   // TANK_CONTROL_1S.PVVX_OUT_DATA.PVVB_DemandsCompleted[10] := False;
   // TANK_CONTROL_1S.PVVX_OUT_DATA.PVVB_DemandsCompleted[9] := False;
   // TANK_CONTROL_1S.PVVX_OUT_DATA.PVVB_DemandsCompleted[8] := False;
   // TANK_CONTROL_1S.PVVX_OUT_DATA.PVVB_DemandsCompleted[7] := False;
   // TANK_CONTROL_1S.PVVX_OUT_DATA.PVVB_DemandsCompleted[6] := False;
   // TANK_CONTROL_1S.PVVX_OUT_DATA.PVVB_DemandsCompleted[5] := False;
   // TANK_CONTROL_6P.DWELL_TIMER.IN := False;
   // TANK_CONTROL_6P.MONITOR_TIMER.IN := False;
   // TANK_CONTROL_6P.ReOx_InitialTargetpHLevelAchieved := False;
   // TANK_CONTROL_1S.PVVX_OUT_DATA.PVVB_DemandsCompleted[4] := False;
   // TANK_CONTROL_1S.PVVX_OUT_DATA.PVVB_DemandsCompleted[3] := False;
   // TANK_CONTROL_1S.PVVX_OUT_DATA.PVVB_DemandsCompleted[2] := False;
   // TANK_CONTROL_1S.PVVX_OUT_DATA.PVVB_DemandsCompleted[1] := False;
   // TANK_CONTROL_1S.PVVX_OUT_DATA.PVVA_Alarms[14] := False;
   // TANK_CONTROL_1S.PVVX_OUT_DATA.PVVA_Alarms[13] := False;
   // TANK_CONTROL_1S.PVVX_OUT_DATA.PVVA_Alarms[12] := False;
   // TANK_CONTROL_1S.PVVX_OUT_DATA.PVVA_Alarms[11] := False;
   // TANK_CONTROL_1S.PVVX_OUT_DATA.PVVA_Alarms[10] := False;
   // TANK_CONTROL_1S.PVVX_OUT_DATA.PVVA_Alarms[9] := False;
   // TANK_CONTROL_1S.PVVX_OUT_DATA.PVVA_Alarms[8] := False;
   // TANK_CONTROL_1S.PVVX_OUT_DATA.PVVA_Alarms[7] := False;
   // TANK_CONTROL_1S.PVVX_OUT_DATA.PVVA_Alarms[6] := False;
   // TANK_CONTROL_1S.PVVX_OUT_DATA.PVVA_Alarms[5] := False;
   // TANK_CONTROL_1S.PVVX_OUT_DATA.PVVA_Alarms[4] := False;
   // TANK_CONTROL_1S.PVVX_OUT_DATA.PVVA_Alarms[3] := False;
   // TANK_CONTROL_1S.PVVX_OUT_DATA.PVVA_Alarms[2] := False;
   // TANK_CONTROL_1S.PVVX_OUT_DATA.PVVA_Alarms[1] := False;
   // TANK_CONTROL_1S.PVVX_OUT_DATA.PVVA_DemandsCompleted[14] := False;
   // TANK_CONTROL_1S.PVVX_OUT_DATA.PVVA_DemandsCompleted[13] := False;
   // TANK_CONTROL_1S.PVVX_OUT_DATA.PVVA_DemandsCompleted[12] := False;
   // TANK_CONTROL_1S.PVVX_OUT_DATA.PVVA_DemandsCompleted[11] := False;
   // TANK_CONTROL_1S.PVVX_OUT_DATA.PVVA_DemandsCompleted[10] := False;
   // TANK_CONTROL_1S.PVVX_OUT_DATA.PVVA_DemandsCompleted[9] := False;
   // TANK_CONTROL_1S.PVVX_OUT_DATA.PVVA_DemandsCompleted[8] := False;
   // TANK_CONTROL_1S.PVVX_OUT_DATA.PVVA_DemandsCompleted[7] := False;
   // TANK_CONTROL_1S.PVVX_OUT_DATA.PVVA_DemandsCompleted[6] := False;
   // TANK_CONTROL_1S.PVVX_OUT_DATA.PVVA_DemandsCompleted[5] := False;
   // TANK_CONTROL_1S.PVVX_OUT_DATA.PVVA_DemandsCompleted[4] := False;
   // TANK_CONTROL_1S.PVVX_OUT_DATA.PVVA_DemandsCompleted[3] := False;
   // TANK_CONTROL_1S.PVVX_OUT_DATA.PVVA_DemandsCompleted[2] := False;
   // TANK_CONTROL_1S.PVVX_OUT_DATA.PVVA_DemandsCompleted[1] := False;
   // TANK_CONTROL_1P.GTT_OUT_DATA.GTT_Alarms[14] := False;
   // TANK_CONTROL_1P.GTT_OUT_DATA.GTT_Alarms[13] := False;
   // TANK_CONTROL_1P.GTT_OUT_DATA.GTT_Alarms[12] := False;
   // TANK_CONTROL_1P.GTT_OUT_DATA.GTT_Alarms[11] := False;
   // TANK_CONTROL_1P.GTT_OUT_DATA.GTT_Alarms[10] := False;
   // TANK_CONTROL_1P.GTT_OUT_DATA.GTT_Alarms[9] := False;
   // TANK_CONTROL_1P.GTT_OUT_DATA.GTT_Alarms[8] := False;
   // TANK_CONTROL_1P.GTT_OUT_DATA.GTT_Alarms[7] := False;
   // TANK_CONTROL_1P.GTT_OUT_DATA.GTT_Alarms[6] := False;
   // TANK_CONTROL_1P.GTT_OUT_DATA.GTT_Alarms[5] := False;
   // TANK_CONTROL_1P.GTT_OUT_DATA.GTT_Alarms[4] := False;
   // TANK_CONTROL_1P.GTT_OUT_DATA.GTT_Alarms[3] := False;
   // TANK_CONTROL_1P.GTT_OUT_DATA.GTT_Alarms[2] := False;
   // TANK_CONTROL_1P.GTT_OUT_DATA.GTT_Alarms[1] := False;
   // TANK_CONTROL_1P.GTT_OUT_DATA.GTT_DemandsCompleted[14] := False;
   // TANK_CONTROL_1P.GTT_OUT_DATA.GTT_DemandsCompleted[13] := False;
   // TANK_CONTROL_1P.GTT_OUT_DATA.GTT_DemandsCompleted[12] := False;
   // TANK_CONTROL_1P.GTT_OUT_DATA.GTT_DemandsCompleted[11] := False;
   // TANK_CONTROL_1P.GTT_OUT_DATA.GTT_DemandsCompleted[10] := False;
   // TANK_CONTROL_1P.GTT_OUT_DATA.GTT_DemandsCompleted[9] := False;
   // TANK_CONTROL_1P.GTT_OUT_DATA.GTT_DemandsCompleted[8] := False;
   // TANK_CONTROL_1P.GTT_OUT_DATA.GTT_DemandsCompleted[7] := False;
   // TANK_CONTROL_1P.GTT_OUT_DATA.GTT_DemandsCompleted[6] := False;
   // TANK_CONTROL_1P.GTT_OUT_DATA.GTT_DemandsCompleted[5] := False;
   // TANK_CONTROL_1P.GTT_OUT_DATA.GTT_DemandsCompleted[4] := False;
   // TANK_CONTROL_1P.GTT_OUT_DATA.GTT_DemandsCompleted[3] := False;
   // TANK_CONTROL_1P.GTT_OUT_DATA.GTT_DemandsCompleted[2] := False;
   // TANK_CONTROL_1P.GTT_OUT_DATA.GTT_DemandsCompleted[1] := False;
   // TANK_CONTROL_1P.PVVX_OUT_DATA.PVVB_Alarms[14] := False;
   // TANK_CONTROL_1P.PVVX_OUT_DATA.PVVB_Alarms[13] := False;
   // TANK_CONTROL_1P.PVVX_OUT_DATA.PVVB_Alarms[12] := False;
   // TANK_CONTROL_1P.PVVX_OUT_DATA.PVVB_Alarms[11] := False;
   // TANK_CONTROL_1P.PVVX_OUT_DATA.PVVB_Alarms[10] := False;
   // TANK_CONTROL_1P.PVVX_OUT_DATA.PVVB_Alarms[9] := False;
   // TANK_CONTROL_1P.PVVX_OUT_DATA.PVVB_Alarms[8] := False;
   // TANK_CONTROL_1P.PVVX_OUT_DATA.PVVB_Alarms[7] := False;
   // TANK_CONTROL_1P.PVVX_OUT_DATA.PVVB_Alarms[6] := False;
   // TANK_CONTROL_1P.PVVX_OUT_DATA.PVVB_Alarms[5] := False;
   // TANK_CONTROL_1P.PVVX_OUT_DATA.PVVB_Alarms[4] := False;
   // TANK_CONTROL_1P.PVVX_OUT_DATA.PVVB_Alarms[3] := False;
   // TANK_CONTROL_1P.PVVX_OUT_DATA.PVVB_Alarms[2] := False;
   // TANK_CONTROL_1P.PVVX_OUT_DATA.PVVB_Alarms[1] := False;
   // TANK_CONTROL_1P.PVVX_OUT_DATA.PVVB_DemandsCompleted[14] := False;
   // TANK_CONTROL_1P.PVVX_OUT_DATA.PVVB_DemandsCompleted[13] := False;
   // TANK_CONTROL_1P.PVVX_OUT_DATA.PVVB_DemandsCompleted[12] := False;
   // TANK_CONTROL_1P.PVVX_OUT_DATA.PVVB_DemandsCompleted[11] := False;
   // TANK_CONTROL_1P.PVVX_OUT_DATA.PVVB_DemandsCompleted[10] := False;
   // TANK_CONTROL_1P.PVVX_OUT_DATA.PVVB_DemandsCompleted[9] := False;
   // TANK_CONTROL_1P.PVVX_OUT_DATA.PVVB_DemandsCompleted[8] := False;
   // TANK_CONTROL_1P.PVVX_OUT_DATA.PVVB_DemandsCompleted[7] := False;
   // TANK_CONTROL_1P.PVVX_OUT_DATA.PVVB_DemandsCompleted[6] := False;
   // TANK_CONTROL_1P.PVVX_OUT_DATA.PVVB_DemandsCompleted[5] := False;
   // TANK_CONTROL_1P.PVVX_OUT_DATA.PVVB_DemandsCompleted[4] := False;
   // TANK_CONTROL_1P.PVVX_OUT_DATA.PVVB_DemandsCompleted[3] := False;
   // TANK_CONTROL_1P.PVVX_OUT_DATA.PVVB_DemandsCompleted[2] := False;
   // TANK_CONTROL_1P.PVVX_OUT_DATA.PVVB_DemandsCompleted[1] := False;
   // TANK_CONTROL_1P.PVVX_OUT_DATA.PVVA_Alarms[14] := False;
   // TANK_CONTROL_1P.PVVX_OUT_DATA.PVVA_Alarms[13] := False;
   // TANK_CONTROL_1P.PVVX_OUT_DATA.PVVA_Alarms[12] := False;
   // TANK_CONTROL_1P.PVVX_OUT_DATA.PVVA_Alarms[11] := False;
   // TANK_CONTROL_1P.PVVX_OUT_DATA.PVVA_Alarms[10] := False;
   // TANK_CONTROL_1P.PVVX_OUT_DATA.PVVA_Alarms[9] := False;
   // TANK_CONTROL_1P.PVVX_OUT_DATA.PVVA_Alarms[8] := False;
   // TANK_CONTROL_1P.PVVX_OUT_DATA.PVVA_Alarms[7] := False;
   // TANK_CONTROL_1P.PVVX_OUT_DATA.PVVA_Alarms[6] := False;
   // TANK_CONTROL_1P.PVVX_OUT_DATA.PVVA_Alarms[5] := False;
   // TANK_CONTROL_1P.PVVX_OUT_DATA.PVVA_Alarms[4] := False;
   // TANK_CONTROL_1P.PVVX_OUT_DATA.PVVA_Alarms[3] := False;
   // TANK_CONTROL_6S.DWELL_TIMER.IN := False;
   // TANK_CONTROL_6S.MONITOR_TIMER.IN := False;
   // TANK_CONTROL_6S.ReOx_InitialTargetpHLevelAchieved := False;
   // TANK_CONTROL_1P.PVVX_OUT_DATA.PVVA_Alarms[2] := False;
   // TANK_CONTROL_1P.PVVX_OUT_DATA.PVVA_Alarms[1] := False;
   // TANK_CONTROL_1P.PVVX_OUT_DATA.PVVA_DemandsCompleted[14] := False;
   // TANK_CONTROL_1P.PVVX_OUT_DATA.PVVA_DemandsCompleted[13] := False;
   // TANK_CONTROL_1P.PVVX_OUT_DATA.PVVA_DemandsCompleted[12] := False;
   // TANK_CONTROL_1P.PVVX_OUT_DATA.PVVA_DemandsCompleted[11] := False;
   // TANK_CONTROL_1P.PVVX_OUT_DATA.PVVA_DemandsCompleted[10] := False;
   // TANK_CONTROL_1P.PVVX_OUT_DATA.PVVA_DemandsCompleted[9] := False;
   // TANK_CONTROL_1P.PVVX_OUT_DATA.PVVA_DemandsCompleted[8] := False;
   // TANK_CONTROL_1P.PVVX_OUT_DATA.PVVA_DemandsCompleted[7] := False;
   // TANK_CONTROL_1P.PVVX_OUT_DATA.PVVA_DemandsCompleted[6] := False;
   // TANK_CONTROL_1P.PVVX_OUT_DATA.PVVA_DemandsCompleted[5] := False;
   // TANK_CONTROL_1P.PVVX_OUT_DATA.PVVA_DemandsCompleted[4] := False;
   // TANK_CONTROL_1P.PVVX_OUT_DATA.PVVA_DemandsCompleted[3] := False;
   // TANK_CONTROL_1P.PVVX_OUT_DATA.PVVA_DemandsCompleted[2] := False;
   // TANK_CONTROL_1P.PVVX_OUT_DATA.PVVA_DemandsCompleted[1] := False;
   // TANK_CONTROL_FPT.GTT_OUT_DATA.GTT_Alarms[14] := False;
   // TANK_CONTROL_FPT.GTT_OUT_DATA.GTT_Alarms[13] := False;
   // TANK_CONTROL_FPT.GTT_OUT_DATA.GTT_Alarms[12] := False;
   // TANK_CONTROL_FPT.GTT_OUT_DATA.GTT_Alarms[11] := False;
   // TANK_CONTROL_FPT.GTT_OUT_DATA.GTT_Alarms[10] := False;
   // TANK_CONTROL_FPT.GTT_OUT_DATA.GTT_Alarms[9] := False;
   // TANK_CONTROL_FPT.GTT_OUT_DATA.GTT_Alarms[8] := False;
   // TANK_CONTROL_FPT.GTT_OUT_DATA.GTT_Alarms[7] := False;
   // TANK_CONTROL_FPT.GTT_OUT_DATA.GTT_Alarms[6] := False;
   // TANK_CONTROL_FPT.GTT_OUT_DATA.GTT_Alarms[5] := False;
   // TANK_CONTROL_FPT.GTT_OUT_DATA.GTT_Alarms[4] := False;
   // TANK_CONTROL_FPT.GTT_OUT_DATA.GTT_Alarms[3] := False;
   // TANK_CONTROL_FPT.GTT_OUT_DATA.GTT_Alarms[2] := False;
   // TANK_CONTROL_FPT.GTT_OUT_DATA.GTT_Alarms[1] := False;
   // TANK_CONTROL_FPT.GTT_OUT_DATA.GTT_DemandsCompleted[14] := False;
   // TANK_CONTROL_FPT.GTT_OUT_DATA.GTT_DemandsCompleted[13] := False;
   // TANK_CONTROL_FPT.GTT_OUT_DATA.GTT_DemandsCompleted[12] := False;
   // TANK_CONTROL_FPT.GTT_OUT_DATA.GTT_DemandsCompleted[11] := False;
   // TANK_CONTROL_FPT.GTT_OUT_DATA.GTT_DemandsCompleted[10] := False;
   // TANK_CONTROL_FPT.GTT_OUT_DATA.GTT_DemandsCompleted[9] := False;
   // TANK_CONTROL_FPT.GTT_OUT_DATA.GTT_DemandsCompleted[8] := False;
   // TANK_CONTROL_FPT.GTT_OUT_DATA.GTT_DemandsCompleted[7] := False;
   // TANK_CONTROL_FPT.GTT_OUT_DATA.GTT_DemandsCompleted[6] := False;
   // TANK_CONTROL_FPT.GTT_OUT_DATA.GTT_DemandsCompleted[5] := False;
   // TANK_CONTROL_FPT.GTT_OUT_DATA.GTT_DemandsCompleted[4] := False;
   // TANK_CONTROL_FPT.GTT_OUT_DATA.GTT_DemandsCompleted[3] := False;
   // TANK_CONTROL_FPT.GTT_OUT_DATA.GTT_DemandsCompleted[2] := False;
   // TANK_CONTROL_FPT.GTT_OUT_DATA.GTT_DemandsCompleted[1] := False;
   // TANK_CONTROL_FPT.PVVX_OUT_DATA.PVVB_Alarms[14] := False;
   // TANK_CONTROL_FPT.PVVX_OUT_DATA.PVVB_Alarms[13] := False;
   // TANK_CONTROL_FPT.PVVX_OUT_DATA.PVVB_Alarms[12] := False;
   // TANK_CONTROL_FPT.PVVX_OUT_DATA.PVVB_Alarms[11] := False;
   // TANK_CONTROL_FPT.PVVX_OUT_DATA.PVVB_Alarms[10] := False;
   // TANK_CONTROL_FPT.PVVX_OUT_DATA.PVVB_Alarms[9] := False;
   // TANK_CONTROL_FPT.PVVX_OUT_DATA.PVVB_Alarms[8] := False;
   // TANK_CONTROL_FPT.PVVX_OUT_DATA.PVVB_Alarms[7] := False;
   // TANK_CONTROL_FPT.PVVX_OUT_DATA.PVVB_Alarms[6] := False;
   // TANK_CONTROL_FPT.PVVX_OUT_DATA.PVVB_Alarms[5] := False;
   // TANK_CONTROL_FPT.PVVX_OUT_DATA.PVVB_Alarms[4] := False;
   // TANK_CONTROL_FPT.PVVX_OUT_DATA.PVVB_Alarms[3] := False;
   // TANK_CONTROL_FPT.PVVX_OUT_DATA.PVVB_Alarms[2] := False;
   // TANK_CONTROL_FPT.PVVX_OUT_DATA.PVVB_Alarms[1] := False;
   // TANK_CONTROL_FPT.PVVX_OUT_DATA.PVVB_DemandsCompleted[14] := False;
   // TANK_CONTROL_FPT.PVVX_OUT_DATA.PVVB_DemandsCompleted[13] := False;
   // TANK_CONTROL_FPT.PVVX_OUT_DATA.PVVB_DemandsCompleted[12] := False;
   // TANK_CONTROL_FPT.PVVX_OUT_DATA.PVVB_DemandsCompleted[11] := False;
   // TANK_CONTROL_FPT.PVVX_OUT_DATA.PVVB_DemandsCompleted[10] := False;
   // TANK_CONTROL_FPT.PVVX_OUT_DATA.PVVB_DemandsCompleted[9] := False;
   // TANK_CONTROL_FPT.PVVX_OUT_DATA.PVVB_DemandsCompleted[8] := False;
   // TANK_CONTROL_FPT.PVVX_OUT_DATA.PVVB_DemandsCompleted[7] := False;
   // TANK_CONTROL_FPT.PVVX_OUT_DATA.PVVB_DemandsCompleted[6] := False;
   // TANK_CONTROL_FPT.PVVX_OUT_DATA.PVVB_DemandsCompleted[5] := False;
   // TANK_CONTROL_FPT.PVVX_OUT_DATA.PVVB_DemandsCompleted[4] := False;
   // TANK_CONTROL_FPT.PVVX_OUT_DATA.PVVB_DemandsCompleted[3] := False;
   // TANK_CONTROL_FPT.PVVX_OUT_DATA.PVVB_DemandsCompleted[2] := False;
   // TANK_CONTROL_FPT.PVVX_OUT_DATA.PVVB_DemandsCompleted[1] := False;
   // TANK_CONTROL_FPT.PVVX_OUT_DATA.PVVA_Alarms[14] := False;
   // TANK_CONTROL_FPT.PVVX_OUT_DATA.PVVA_Alarms[13] := False;
   // TANK_CONTROL_FPT.PVVX_OUT_DATA.PVVA_Alarms[12] := False;
   // TANK_CONTROL_FPT.PVVX_OUT_DATA.PVVA_Alarms[11] := False;
   // TANK_CONTROL_FPT.PVVX_OUT_DATA.PVVA_Alarms[10] := False;
   // TANK_CONTROL_FPT.PVVX_OUT_DATA.PVVA_Alarms[9] := False;
   // TANK_CONTROL_FPT.PVVX_OUT_DATA.PVVA_Alarms[8] := False;
   // TANK_CONTROL_FPT.PVVX_OUT_DATA.PVVA_Alarms[7] := False;
   // TANK_CONTROL_FPT.PVVX_OUT_DATA.PVVA_Alarms[6] := False;
   // TANK_CONTROL_FPT.PVVX_OUT_DATA.PVVA_Alarms[5] := False;
   // TANK_CONTROL_FPT.PVVX_OUT_DATA.PVVA_Alarms[4] := False;
   // TANK_CONTROL_FPT.PVVX_OUT_DATA.PVVA_Alarms[3] := False;
   // TANK_CONTROL_FPT.PVVX_OUT_DATA.PVVA_Alarms[2] := False;
   // TANK_CONTROL_FPT.PVVX_OUT_DATA.PVVA_Alarms[1] := False;
   // TANK_CONTROL_FPT.PVVX_OUT_DATA.PVVA_DemandsCompleted[14] := False;
   // TANK_CONTROL_FPT.PVVX_OUT_DATA.PVVA_DemandsCompleted[13] := False;
   // TANK_CONTROL_FPT.PVVX_OUT_DATA.PVVA_DemandsCompleted[12] := False;
   // TANK_CONTROL_FPT.PVVX_OUT_DATA.PVVA_DemandsCompleted[11] := False;
   // TANK_CONTROL_FPT.PVVX_OUT_DATA.PVVA_DemandsCompleted[10] := False;
   // TANK_CONTROL_FPT.PVVX_OUT_DATA.PVVA_DemandsCompleted[9] := False;
   // TANK_CONTROL_FPT.PVVX_OUT_DATA.PVVA_DemandsCompleted[8] := False;
   // TANK_CONTROL_FPT.PVVX_OUT_DATA.PVVA_DemandsCompleted[7] := False;
   // TANK_CONTROL_FPT.PVVX_OUT_DATA.PVVA_DemandsCompleted[6] := False;
   // TANK_CONTROL_FPT.PVVX_OUT_DATA.PVVA_DemandsCompleted[5] := False;
   // TANK_CONTROL_FPT.PVVX_OUT_DATA.PVVA_DemandsCompleted[4] := False;
   // TANK_CONTROL_FPT.PVVX_OUT_DATA.PVVA_DemandsCompleted[3] := False;
   // TANK_CONTROL_FPT.PVVX_OUT_DATA.PVVA_DemandsCompleted[2] := False;
   // TANK_CONTROL_FPT.PVVX_OUT_DATA.PVVA_DemandsCompleted[1] := False;
   // TANK_CONTROL_APT.DWELL_TIMER.IN := False;
   // TANK_CONTROL_APT.MONITOR_TIMER.IN := False;
   // TANK_CONTROL_APT.ReOx_InitialTargetpHLevelAchieved := False;
   // DWELL_TIMER.IN := False;
   // XEOX_TIMER.IN := False;
   // XEOX_PAUSE_TIMER.IN := False;
BEGIN
   // Reset HMI Warnings. These will be re-enabled on a scan-cycle if the HMI Warning is intended to persist.
   "1092_HMI_OP_FLAGS".HMI_Warnings.Active := False;
   // Set the start button to false by default, only set it true under state init, and under correct conditions.
   "1092_HMI_OP_FLAGS".StartButtonEnabled := False;
   IF #State.System <> #State_Shutdown THEN
       // Keep the shutdown reset flag high if not in a reset state.
       #ShutdownStageReset := true;
       // Let GCU know we're not in a shutdown state
       "58_INTRNL_COMMS".BWT_TO_GCU.SHT_DN := False;
   END_IF;
   // If the HMI has signalled to stop treatment, or GCU has shutdown, also shut down BWTS.
   IF "1090_HMI_IP_FLAGS".StopTreatment OR "58_INTRNL_COMMS".GCU_TO_BWT.SHT_DN THEN
       #State.System := #State_Shutdown;
   END_IF;

   (* 
       Main case structure #State.System:
       This main case structure dictates the major phases that group tanks together.
       The system state constrains the state which each tank can be in at any one time.
       The naming convention for each system state is based on the major system events
       take place within the state. The tank states can be descirbed as follows:
       #State_Init: The tanks may only be in Init state.
       #State_PreDwell: The tanks may only bein Pre-Dwell state.
       #State_DeOx: The tanks may only bein Pre-Dwell, DeOx, or Mid-Dwell states.
       #State_DwellAndReOx: The tanks may only be in Mid-Dwell, ReOx, or Post-Dwell states.
       #State_DwellAndComplete: The tanks may only bein Post-Dwell or Done states.
   *)
   CASE #State.System OF
       #State_Init:
           (* 
               Waiting for start signal, Continue to populate the system data such as 
               calculations of treamtnet time, and IGG warning times until user selects start
           *)
           "1131_CALC_HEALTHY_TANKS"();
           "1132_CALC_ACTIVE_TANKS"();
           "58_INTRNL_COMMS".BWT_TO_GCU.SPLY_GAS := False;
           "58_INTRNL_COMMS".BWT_TO_GCU.STP_GAS := True;
           "58_INTRNL_COMMS".BWT_TO_GCU.PREP_GAS := False;
           "1191_SYSTEM_VARIABLES".TreatmentTime := "1130_CALC_TREATMENT_TIME"();
           "1191_SYSTEM_VARIABLES".StartIGGWarningsTime := ("1096_ADJUSTABLE_CONSTANTS".VoyageTime - "1191_SYSTEM_VARIABLES".TreatmentTime + "1190_FIXED_CONSTANTS".PreDwell_Time - LT#2h);
           FOR #Index := 1 TO #NumberOfTanks DO
               #TankData[#Index].TankState := #TankState_Init;
           END_FOR;
           // Push warning flag if the voyage time is less than the calculated treatment time.
           IF "1096_ADJUSTABLE_CONSTANTS".VoyageTime < "1191_SYSTEM_VARIABLES".TreatmentTime THEN
               "1092_HMI_OP_FLAGS".VoyageLessThanTreatmentTime := True;
           ELSE
               "1092_HMI_OP_FLAGS".VoyageLessThanTreatmentTime := False;
           END_IF;
           IF NOT ("1092_HMI_OP_FLAGS".VoyageLessThanTreatmentTime) AND NOT ("1092_HMI_OP_FLAGS".NoTanksActive) THEN
               "1092_HMI_OP_FLAGS".StartButtonEnabled := True;
           END_IF;
           (* 
               User has pushed the start treatment button, set the BWT process to start
               by moving the tanks into a pre-dwell state and starting the timers. Call all
               appropriate resets to provide a clean new environment for this process 
           *)
           IF "1090_HMI_IP_FLAGS".StartTreatment THEN
               // populate tank data for initialization.
               FOR #Index := 1 TO #NumberOfTanks DO
                   #TankData[#Index].TankState := #TankState_PreDwell;
                   #TankData[#Index].TankID := #Index;
                   #TankData[#Index].Active := "1096_ADJUSTABLE_CONSTANTS".TankIDActive[#Index];
               END_FOR;
               // Set system state to predwell for next cycle
               #State.System := #State_PreDwell;
               // Reset the dwell timer.
               #DWELL_TIMER(IN := False,
                            PT := #MaxTimerPT,
                            R := True);
               // Reset the ReOx/DeOx timer.
               #XEOX_TIMER(IN := False,
                           PT := #MaxTimerPT,
                           R := True);
               // Reset the ReOx/DeOx pause timer.
               #XEOX_PAUSE_TIMER(IN := False,
                                 PT := #MaxTimerPT,
                                 R := True);
           END_IF;
       #State_PreDwell:
           #DWELL_TIMER(IN := True,
                        PT := #MaxTimerPT,
                        R := False);
           // Check The IGG Warning timers (BWMS-072)
           // Check FOR IGG Warnings based on current Pre Dwell Time.
           IF #DWELL_TIMER.ET >= "1191_SYSTEM_VARIABLES".StartIGGWarningsTime THEN
               "1092_HMI_OP_FLAGS".HMI_Warnings.Active := True;
               "1092_HMI_OP_FLAGS".HMI_Warnings.Message := 'Start IGG 60 Minute Warning';
           ELSIF #DWELL_TIMER.ET >= ("1191_SYSTEM_VARIABLES".StartIGGWarningsTime + LT#15m) THEN
               "1092_HMI_OP_FLAGS".HMI_Warnings.Active := True;
               "1092_HMI_OP_FLAGS".HMI_Warnings.Message := 'Start IGG 45 Minute Warning';
           ELSIF #DWELL_TIMER.ET >= ("1191_SYSTEM_VARIABLES".StartIGGWarningsTime + LT#30m) THEN
               "1092_HMI_OP_FLAGS".HMI_Warnings.Active := True;
               "1092_HMI_OP_FLAGS".HMI_Warnings.Message := 'Start IGG 30 Minute Warning';
           ELSIF #DWELL_TIMER.ET >= ("1191_SYSTEM_VARIABLES".StartIGGWarningsTime + LT#45m) THEN
               "1092_HMI_OP_FLAGS".HMI_Warnings.Active := True;
               "1092_HMI_OP_FLAGS".HMI_Warnings.Message := 'Start IGG 15 Minute Warning';
           ELSIF #DWELL_TIMER.ET >= ("1191_SYSTEM_VARIABLES".StartIGGWarningsTime + LT#60m) THEN
               "1092_HMI_OP_FLAGS".HMI_Warnings.Active := True;
               "1092_HMI_OP_FLAGS".HMI_Warnings.Message := 'Start IGG - Operator Confirmation';
           ELSE
               "1092_HMI_OP_FLAGS".HMI_Warnings.Active := False;
               "1092_HMI_OP_FLAGS".HMI_Warnings.Message := '';
           END_IF;

           // Pre-dwell timer has elapsed, sufficient voyage time has occured for BWT to start, IG is ready. GCU is ready.
           IF ("1191_SYSTEM_VARIABLES".FromIGG_InertGasReady AND "58_INTRNL_COMMS".GCU_TO_BWT.GAS_AVLBL
               AND #DWELL_TIMER.ET >= ("1096_ADJUSTABLE_CONSTANTS".VoyageTime - "1191_SYSTEM_VARIABLES".TreatmentTime + "1190_FIXED_CONSTANTS".PreDwell_Time)) THEN
               // Reset the supply to deck stage to zero, move state to deox & supply to deck
               #DECK_MANAGE_START_SUPPLY.Stage := 0;
               #State.System := #State_DeOx;
               #State.DeOx := #State_DeOx_SupplyToDeck;
           END_IF;

       #State_DeOx:
           CASE #State.DeOx OF
               #State_DeOx_SupplyToDeck:
                   IF #DECK_MANAGE_START_SUPPLY.ShutdownDemand THEN
                       // Deck supply has failed, shutdown demand.
                       #State.System := #State_Shutdown;
                   ELSIF "1092_HMI_OP_FLAGS".DeckSupplyOk THEN
                       // Deck supply is established, start DeOxygenation on treatment group 1.
                       #State.TreatmentGroup := 1;
                       #State.DeOx := #State_DeOx_ClosePVV;
                   ELSE
                       // Deck supply is not complete yet, run supply to deck automation.
                       #DECK_MANAGE_START_SUPPLY();
                       "58_INTRNL_COMMS".BWT_TO_GCU.SPLY_GAS := True;
                       "58_INTRNL_COMMS".BWT_TO_GCU.STP_GAS := False;
                   END_IF;
               #State_DeOx_ClosePVV:
                   // Does this setup use PVV? If so, no electronic actuation is required, jump to openGTTs.
                   IF "1090_HMI_IP_FLAGS".PressVacuumValves THEN
                       #State.DeOx := #State_DeOx_OpenGTT;
                   ELSE
                       // Check if ready to move to to openning GTTs once appropriate PVVs have reported demand completion.
                       #NextStageCheck := "1151_NEXT_STAGE_CHECK_PVV"(AlarmState := #State_Shutdown, PVVX_OUT := #PVVX_OUT, State := #State, TankData := #TankData);
                       IF #NextStageCheck.Demand_Complete AND NOT #NextStageCheck.Alarm_Active THEN
                           #State.DeOx := #State_DeOx_OpenGTT;
                       END_IF;
                   END_IF;
               #State_DeOx_OpenGTT:
                   // Check if ready to move to monitoring stage once appropriate GTTs have reported demand completion.
                   #NextStageCheck := "1150_NEXT_STAGE_CHECK_GTT"(AlarmState := #State_Shutdown, GTT_OUT := #GTT_OUT, State := #State, TankData := #TankData);
                   IF #NextStageCheck.Demand_Complete AND NOT #NextStageCheck.Alarm_Active THEN
                       // Reset timer information for this new treatment group
                       #XEOX_PausedTime := LT#0s;
                       #XEOX_TIMER(IN := False,
                                   PT := "1190_FIXED_CONSTANTS".DeOxMin_Time + #XEOX_PausedTime,
                                   R := True);
                       #XEOX_PAUSE_TIMER(IN := False,
                                         PT := "1190_FIXED_CONSTANTS".MaxDOPause_Time,
                                         R := True);
                       #State.DeOx := #State_DeOx_Monitor;
                       "1134_MOVE_TANKS_INGROUP_NEW_STATE"(TankData := #TankData,
                                                          State := #State,
                                                          NewState := #TankState_DeOx);
                   END_IF;
               #State_DeOx_Monitor:
                   // Has DeOxygenation completed? If so, close GTTs if this is not the last treatment group.
                   // If this is the last treatment group, stop the supply to deck first (then close GTTs) to avoid
                   // pressure build up on the main deck line.
                   IF #XEOX_TIMER.Q THEN
                       #NextStageCheck := "1153_NEXT_STAGE_CHECK_XEOX"(AlarmState := #State_Shutdown, State := #State, TankData := #TankData);
                       IF #NextStageCheck.Demand_Complete AND NOT #NextStageCheck.Alarm_Active THEN
                           #NextTreatmentGroup := "1136_CALC_NEXT_TREATMENT_GROUP"(NumberOfTreatmentGroups := "1190_FIXED_CONSTANTS".NumberOfTreatmentGroups, State := #State, TankData := #TankData);
                           IF #NextTreatmentGroup = -1 THEN
                               #DECK_MANAGE_STOP_SUPPLY.Stage := 0;
                               #State.DeOx := #State_DeOx_StopSupplyToDeck;
                           ELSE
                               #State.DeOx := #State_DeOx_CloseGTT;
                           END_IF;
                       END_IF;
                   ELSE
                       IF "1191_SYSTEM_VARIABLES".FromIGG_InertGasReady AND "58_INTRNL_COMMS".GCU_TO_BWT.GAS_AVLBL THEN
                           // continue counting on the deox timer as GCU & IG are in healthy states.
                           // increment the paused time as this shall be added to the deoxmin_time due to stoppage.
                           #XEOX_PausedTime += #XEOX_PAUSE_TIMER.ET;
                           #XEOX_TIMER(IN := True,
                                       PT := "1190_FIXED_CONSTANTS".DeOxMin_Time + #XEOX_PausedTime,
                                       R := False);
                           // keep Dissoloved Oxygen pause timer in reset state.
                           #XEOX_PAUSE_TIMER(IN := False,
                                             PT := "1190_FIXED_CONSTANTS".MaxDOPause_Time,
                                             R := True);
                       ELSE
                           // there is a problem with the IG and/or GCU: increment the pause timer, the maximum
                           // DO pause time shall cause a halt of the BWT Process.
                           IF #XEOX_PAUSE_TIMER.Q THEN
                               // Halt BWT Process (tbd in BMWS-098)
                               #State.System := #State_Shutdown;
                           ELSE
                               // Keep deox timer paused, whilst pause timer increments.
                               #XEOX_TIMER(IN := False,
                                           PT := "1190_FIXED_CONSTANTS".DeOxMin_Time,
                                           R := False);
                               #XEOX_PAUSE_TIMER(IN := True,
                                                 PT := "1190_FIXED_CONSTANTS".MaxDOPause_Time,
                                                 R := False);
                           END_IF;
                       END_IF;
                   END_IF;
               #State_DeOx_CloseGTT:
                   // Check if ready to move to mid-dwell stage once appropriate GTTs have reported demand completion
                   #NextStageCheck := "1150_NEXT_STAGE_CHECK_GTT"(AlarmState := #State_Shutdown, GTT_OUT := #GTT_OUT, State := #State, TankData := #TankData);
                   IF #NextStageCheck.Demand_Complete AND NOT #NextStageCheck.Alarm_Active THEN
                       // All tanks in this treatment group are now de-oxed, move them to mid-dwell tank state.
                       "1134_MOVE_TANKS_INGROUP_NEW_STATE"(TankData := #TankData,
                                                          State := #State,
                                                          NewState := #TankState_MidDwell);
                       // If this is the last treatment group. If this is not the last treatment group,
                       // is the system ready to restart on the next treatment group in order?
                      #NextTreatmentGroup := "1136_CALC_NEXT_TREATMENT_GROUP"(NumberOfTreatmentGroups := "1190_FIXED_CONSTANTS".NumberOfTreatmentGroups, State := #State, TankData := #TankData);
                       IF #NextTreatmentGroup = -1 THEN
                           #State.TreatmentGroup := 1;
                           #State.System := #State_DwellAndReOx;
                           #State.ReOx := #State_DwellAndReOx_WaitMidDwell;
                       ELSE
                           #State.TreatmentGroup := #NextTreatmentGroup;
                           #State.DeOx := #State_DeOx_ClosePVV;
                       END_IF;
                   END_IF;
               #State_DeOx_StopSupplyToDeck:
                   IF #DECK_MANAGE_STOP_SUPPLY.ShutdownDemand THEN
                       // Deck supply has failed, shutdown demand.
                       #State.System := #State_Shutdown;
                   ELSIF #DECK_MANAGE_STOP_SUPPLY.StopDeckSupplyDone THEN
                       // Deck stop supply is complete, close the final set of GTT valves.
                       #State.DeOx := #State_DeOx_CloseGTT;
                   ELSE
                       // Deck stop supply is not complete yet, run stop supply to deck automation.
                       #DECK_MANAGE_STOP_SUPPLY();
                       "58_INTRNL_COMMS".BWT_TO_GCU.SPLY_GAS := False;
                       "58_INTRNL_COMMS".BWT_TO_GCU.STP_GAS := True;
                   END_IF;
           END_CASE;

       #State_DwellAndReOx:
           CASE #State.ReOx OF
               #State_DwellAndReOx_WaitMidDwell:
                   #NextStageCheck := "1152_NEXT_STAGE_CHECK_TIMER"(AlarmState := #State_Shutdown, State := #State, TankData := #TankData);
                   IF #NextStageCheck.Demand_Complete AND NOT #NextStageCheck.Alarm_Active THEN
                       "1134_MOVE_TANKS_INGROUP_NEW_STATE"(TankData := #TankData,
                                                          State := #State,
                                                          NewState := #TankState_ReOx);
                       // If this is the first treatment group to finish mid-dwell, open the supply to deck, then open PVV.
                       // Else, jump directly to the open PVV stage as the supply to deck will already be established.
                       IF #State.TreatmentGroup = 1 THEN
                           // Start deck supply starts with the first treatment group to have finished mid-dwell (BWMS-131)
                           #DECK_MANAGE_START_SUPPLY.Stage := 0;
                           "58_INTRNL_COMMS".BWT_TO_GCU.SPLY_GAS := True;
                           "58_INTRNL_COMMS".BWT_TO_GCU.STP_GAS := False;
                           #State.ReOx := #State_DwellAndReOx_SupplyToDeck;
                       ELSE
                           #State.ReOx := #State_DwellAndReOx_OpenPVV;
                       END_IF;
                   END_IF;

                   IF #State.TreatmentGroup = 1 THEN
                       IF "1191_SYSTEM_VARIABLES".MidDwell_ElapsedTime >= "1190_FIXED_CONSTANTS".MidDwell_Time - LT#1h THEN
                           // BWMS-127: Warn of re-oxygenation starting in 1h.
                           "1092_HMI_OP_FLAGS".HMI_Warnings.Active := True;
                           "1092_HMI_OP_FLAGS".HMI_Warnings.Message := 'Re-Oxygenation will begin in 1 hour. Switch on additional generator power for this process as required';
                       ELSIF "1191_SYSTEM_VARIABLES".MidDwell_ElapsedTime >= "1190_FIXED_CONSTANTS".MidDwell_Time - LT#30m THEN
                           // BWMS-128: Start the GCU Process here
                           "58_INTRNL_COMMS".BWT_TO_GCU.PREP_GAS := True;
                       END_IF;
                   END_IF;

                   // NOTE: SHOULD THERE BE AN ADDITIONAL 2h TON HERE TO MAKE SURE A DWELL PERIOD IS SUFFICIENT?
                   // Currently: if there is a sufficient number of treatment groups there is a possiblity that TG1 will have completed mid-dwell
                   // as the system transition into mid-dwell and will therefre want to start the ReOx gas supply immediately after the final TG has 
                   // completed DeOx.